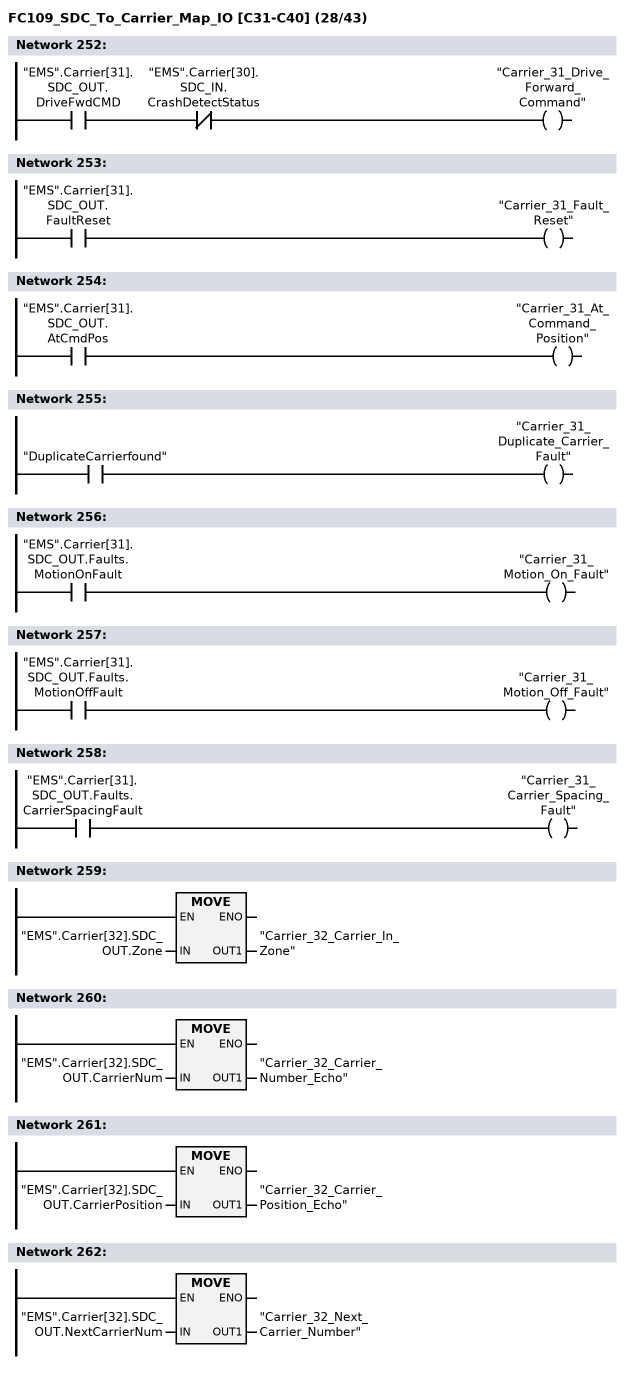
   RUNG wire#powerrail
      Contact( "EMS".Carrier[31].SDC_OUT.DriveFwdCMD )
      I_Contact( "EMS".Carrier[30].SDC_IN.CrashDetectStatus )
      Coil( "Carrier_31_Drive_Forward_Command" )
   END_RUNG
   // the same network as SCL:
   "Carrier_31_Drive_Forward_Command" := "EMS".Carrier[31].SDC_OUT.DriveFwdCMD AND NOT "EMS".Carrier[30].SDC_IN.CrashDetectStatus;
END_REGION

REGION Network 253
   RUNG wire#powerrail
      Contact( "EMS".Carrier[31].SDC_OUT.FaultReset )
      Coil( "Carrier_31_Fault_Reset" )
   END_RUNG
   // the same network as SCL:
   "Carrier_31_Fault_Reset" := "EMS".Carrier[31].SDC_OUT.FaultReset;
END_REGION

REGION Network 254
   RUNG wire#powerrail
      Contact( "EMS".Carrier[31].SDC_OUT.AtCmdPos )
      Coil( "Carrier_31_At_Command_Position" )
   END_RUNG
   // the same network as SCL:
   "Carrier_31_At_Command_Position" := "EMS".Carrier[31].SDC_OUT.AtCmdPos;
END_REGION

REGION Network 255
   RUNG wire#powerrail
      Contact( "DuplicateCarrierfound" )
      Coil( "Carrier_31_Duplicate_Carrier_Fault" )
   END_RUNG
   // the same network as SCL:
   "Carrier_31_Duplicate_Carrier_Fault" := "DuplicateCarrierfound";
END_REGION

REGION Network 256
   RUNG wire#powerrail
      Contact( "EMS".Carrier[31].SDC_OUT.Faults.MotionOnFault )
      Coil( "Carrier_31_Motion_On_Fault" )
   END_RUNG
   // the same network as SCL:
   "Carrier_31_Motion_On_Fault" := "EMS".Carrier[31].SDC_OUT.Faults.MotionOnFault;
END_REGION

REGION Network 257
   RUNG wire#powerrail
      Contact( "EMS".Carrier[31].SDC_OUT.Faults.MotionOffFault )
      Coil( "Carrier_31_Motion_Off_Fault" )
   END_RUNG
   // the same network as SCL:
   "Carrier_31_Motion_Off_Fault" := "EMS".Carrier[31].SDC_OUT.Faults.MotionOffFault;
END_REGION

REGION Network 258
   RUNG wire#powerrail
      Contact( "EMS".Carrier[31].SDC_OUT.Faults.CarrierSpacingFault )
      Coil( "Carrier_31_Carrier_Spacing_Fault" )
   END_RUNG
   // the same network as SCL:
   "Carrier_31_Carrier_Spacing_Fault" := "EMS".Carrier[31].SDC_OUT.Faults.CarrierSpacingFault;
END_REGION

REGION Network 259
   RUNG wire#powerrail
      Move(in := "EMS".Carrier[32].SDC_OUT.Zone, out1 => "Carrier_32_Carrier_In_Zone")
   END_RUNG
   // the same network as SCL:
   "Carrier_32_Carrier_In_Zone" := "EMS".Carrier[32].SDC_OUT.Zone;
END_REGION

REGION Network 260
   RUNG wire#powerrail
      Move(in := "EMS".Carrier[32].SDC_OUT.CarrierNum, out1 => "Carrier_32_Carrier_Number_Echo")
   END_RUNG
   // the same network as SCL:
   "Carrier_32_Carrier_Number_Echo" := "EMS".Carrier[32].SDC_OUT.CarrierNum;
END_REGION

REGION Network 261
   RUNG wire#powerrail
      Move(in := "EMS".Carrier[32].SDC_OUT.CarrierPosition, out1 => "Carrier_32_Carrier_Position_Echo")
   END_RUNG
   // the same network as SCL:
   "Carrier_32_Carrier_Position_Echo" := "EMS".Carrier[32].SDC_OUT.CarrierPosition;
END_REGION

REGION Network 262
   RUNG wire#powerrail
      Move(in := "EMS".Carrier[32].SDC_OUT.NextCarrierNum, out1 => "Carrier_32_Next_Carrier_Number")
   END_RUNG
   // the same network as SCL:
   "Carrier_32_Next_Carrier_Number" := "EMS".Carrier[32].SDC_OUT.NextCarrierNum;
END_REGION

REGION Network 263
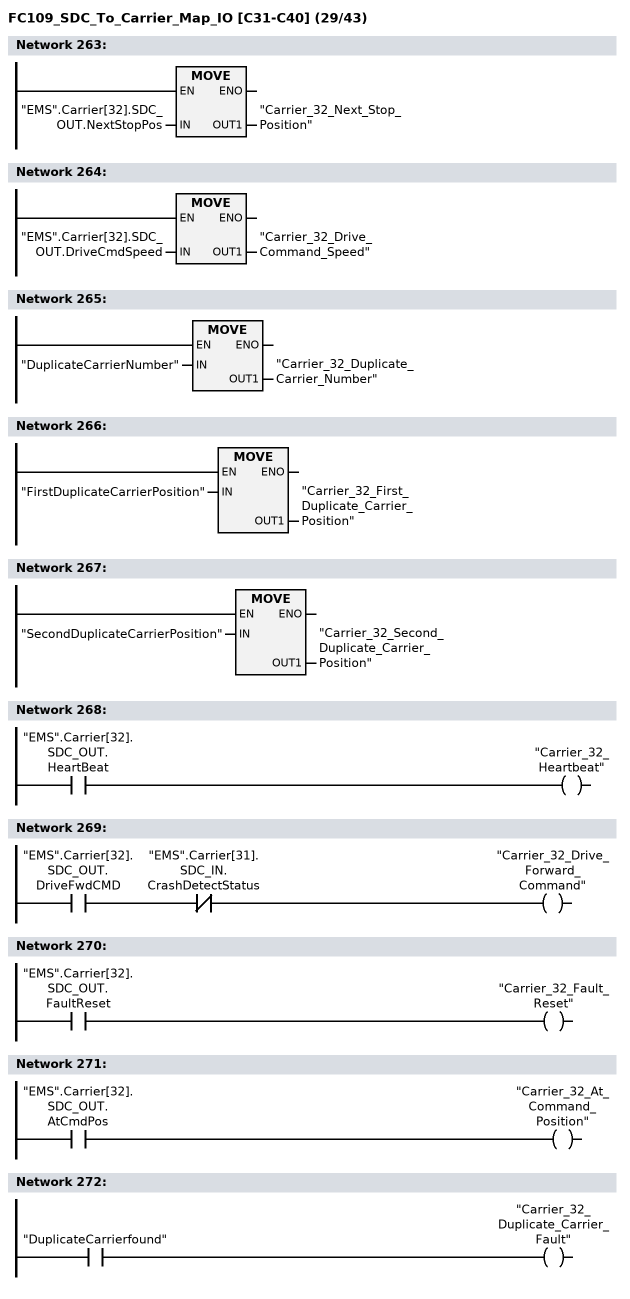
   RUNG wire#powerrail
      Move(in := "EMS".Carrier[32].SDC_OUT.NextStopPos, out1 => "Carrier_32_Next_Stop_Position")
   END_RUNG
   // the same network as SCL:
   "Carrier_32_Next_Stop_Position" := "EMS".Carrier[32].SDC_OUT.NextStopPos;
END_REGION

REGION Network 264
   RUNG wire#powerrail
      Move(in := "EMS".Carrier[32].SDC_OUT.DriveCmdSpeed, out1 => "Carrier_32_Drive_Command_Speed")
   END_RUNG
   // the same network as SCL:
   "Carrier_32_Drive_Command_Speed" := "EMS".Carrier[32].SDC_OUT.DriveCmdSpeed;
END_REGION

REGION Network 265
   RUNG wire#powerrail
      Move(in := "DuplicateCarrierNumber", out1 => "Carrier_32_Duplicate_Carrier_Number")
   END_RUNG
   // the same network as SCL:
   "Carrier_32_Duplicate_Carrier_Number" := "DuplicateCarrierNumber";
END_REGION

REGION Network 266
   RUNG wire#powerrail
      Move(in := "FirstDuplicateCarrierPosition", out1 => "Carrier_32_First_Duplicate_Carrier_Position")
   END_RUNG
   // the same network as SCL:
   "Carrier_32_First_Duplicate_Carrier_Position" := "FirstDuplicateCarrierPosition";
END_REGION

REGION Network 267
   RUNG wire#powerrail
      Move(in := "SecondDuplicateCarrierPosition", out1 => "Carrier_32_Second_Duplicate_Carrier_Position")
   END_RUNG
   // the same network as SCL:
   "Carrier_32_Second_Duplicate_Carrier_Position" := "SecondDuplicateCarrierPosition";
END_REGION

REGION Network 268
   RUNG wire#powerrail
      Contact( "EMS".Carrier[32].SDC_OUT.HeartBeat )
      Coil( "Carrier_32_Heartbeat" )
   END_RUNG
   // the same network as SCL:
   "Carrier_32_Heartbeat" := "EMS".Carrier[32].SDC_OUT.HeartBeat;
END_REGION

REGION Network 269
   RUNG wire#powerrail
      Contact( "EMS".Carrier[32].SDC_OUT.DriveFwdCMD )
      I_Contact( "EMS".Carrier[31].SDC_IN.CrashDetectStatus )
      Coil( "Carrier_32_Drive_Forward_Command" )
   END_RUNG
   // the same network as SCL:
   "Carrier_32_Drive_Forward_Command" := "EMS".Carrier[32].SDC_OUT.DriveFwdCMD AND NOT "EMS".Carrier[31].SDC_IN.CrashDetectStatus;
END_REGION

REGION Network 270
   RUNG wire#powerrail
      Contact( "EMS".Carrier[32].SDC_OUT.FaultReset )
      Coil( "Carrier_32_Fault_Reset" )
   END_RUNG
   // the same network as SCL:
   "Carrier_32_Fault_Reset" := "EMS".Carrier[32].SDC_OUT.FaultReset;
END_REGION

REGION Network 271
   RUNG wire#powerrail
      Contact( "EMS".Carrier[32].SDC_OUT.AtCmdPos )
      Coil( "Carrier_32_At_Command_Position" )
   END_RUNG
   // the same network as SCL:
   "Carrier_32_At_Command_Position" := "EMS".Carrier[32].SDC_OUT.AtCmdPos;
END_REGION

REGION Network 272
   RUNG wire#powerrail
      Contact( "DuplicateCarrierfound" )
      Coil( "Carrier_32_Duplicate_Carrier_Fault" )
   END_RUNG
   // the same network as SCL:
   "Carrier_32_Duplicate_Carrier_Fault" := "DuplicateCarrierfound";
END_REGION

REGION Network 273
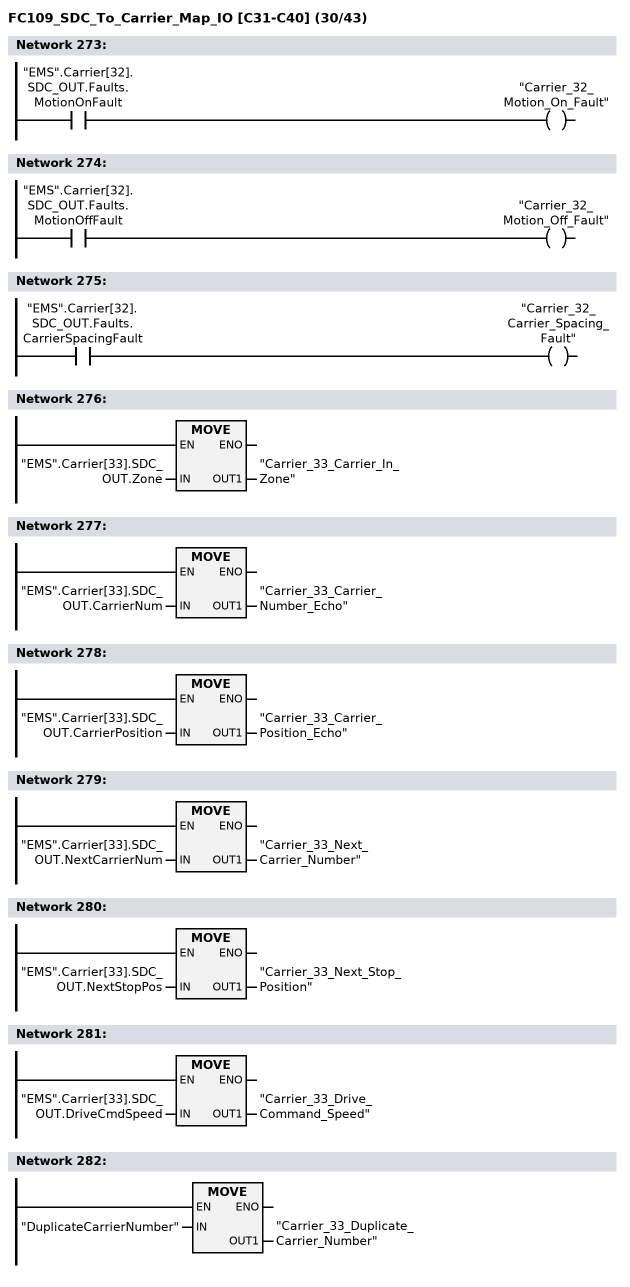
   RUNG wire#powerrail
      Contact( "EMS".Carrier[32].SDC_OUT.Faults.MotionOnFault )
      Coil( "Carrier_32_Motion_On_Fault" )
   END_RUNG
   // the same network as SCL:
   "Carrier_32_Motion_On_Fault" := "EMS".Carrier[32].SDC_OUT.Faults.MotionOnFault;
END_REGION

REGION Network 274
   RUNG wire#powerrail
      Contact( "EMS".Carrier[32].SDC_OUT.Faults.MotionOffFault )
      Coil( "Carrier_32_Motion_Off_Fault" )
   END_RUNG
   // the same network as SCL:
   "Carrier_32_Motion_Off_Fault" := "EMS".Carrier[32].SDC_OUT.Faults.MotionOffFault;
END_REGION

REGION Network 275
   RUNG wire#powerrail
      Contact( "EMS".Carrier[32].SDC_OUT.Faults.CarrierSpacingFault )
      Coil( "Carrier_32_Carrier_Spacing_Fault" )
   END_RUNG
   // the same network as SCL:
   "Carrier_32_Carrier_Spacing_Fault" := "EMS".Carrier[32].SDC_OUT.Faults.CarrierSpacingFault;
END_REGION

REGION Network 276
   RUNG wire#powerrail
      Move(in := "EMS".Carrier[33].SDC_OUT.Zone, out1 => "Carrier_33_Carrier_In_Zone")
   END_RUNG
   // the same network as SCL:
   "Carrier_33_Carrier_In_Zone" := "EMS".Carrier[33].SDC_OUT.Zone;
END_REGION

REGION Network 277
   RUNG wire#powerrail
      Move(in := "EMS".Carrier[33].SDC_OUT.CarrierNum, out1 => "Carrier_33_Carrier_Number_Echo")
   END_RUNG
   // the same network as SCL:
   "Carrier_33_Carrier_Number_Echo" := "EMS".Carrier[33].SDC_OUT.CarrierNum;
END_REGION

REGION Network 278
   RUNG wire#powerrail
      Move(in := "EMS".Carrier[33].SDC_OUT.CarrierPosition, out1 => "Carrier_33_Carrier_Position_Echo")
   END_RUNG
   // the same network as SCL:
   "Carrier_33_Carrier_Position_Echo" := "EMS".Carrier[33].SDC_OUT.CarrierPosition;
END_REGION

REGION Network 279
   RUNG wire#powerrail
      Move(in := "EMS".Carrier[33].SDC_OUT.NextCarrierNum, out1 => "Carrier_33_Next_Carrier_Number")
   END_RUNG
   // the same network as SCL:
   "Carrier_33_Next_Carrier_Number" := "EMS".Carrier[33].SDC_OUT.NextCarrierNum;
END_REGION

REGION Network 280
   RUNG wire#powerrail
      Move(in := "EMS".Carrier[33].SDC_OUT.NextStopPos, out1 => "Carrier_33_Next_Stop_Position")
   END_RUNG
   // the same network as SCL:
   "Carrier_33_Next_Stop_Position" := "EMS".Carrier[33].SDC_OUT.NextStopPos;
END_REGION

REGION Network 281
   RUNG wire#powerrail
      Move(in := "EMS".Carrier[33].SDC_OUT.DriveCmdSpeed, out1 => "Carrier_33_Drive_Command_Speed")
   END_RUNG
   // the same network as SCL:
   "Carrier_33_Drive_Command_Speed" := "EMS".Carrier[33].SDC_OUT.DriveCmdSpeed;
END_REGION

REGION Network 282
   RUNG wire#powerrail
      Move(in := "DuplicateCarrierNumber", out1 => "Carrier_33_Duplicate_Carrier_Number")
   END_RUNG
   // the same network as SCL:
   "Carrier_33_Duplicate_Carrier_Number" := "DuplicateCarrierNumber";
END_REGION

REGION Network 283
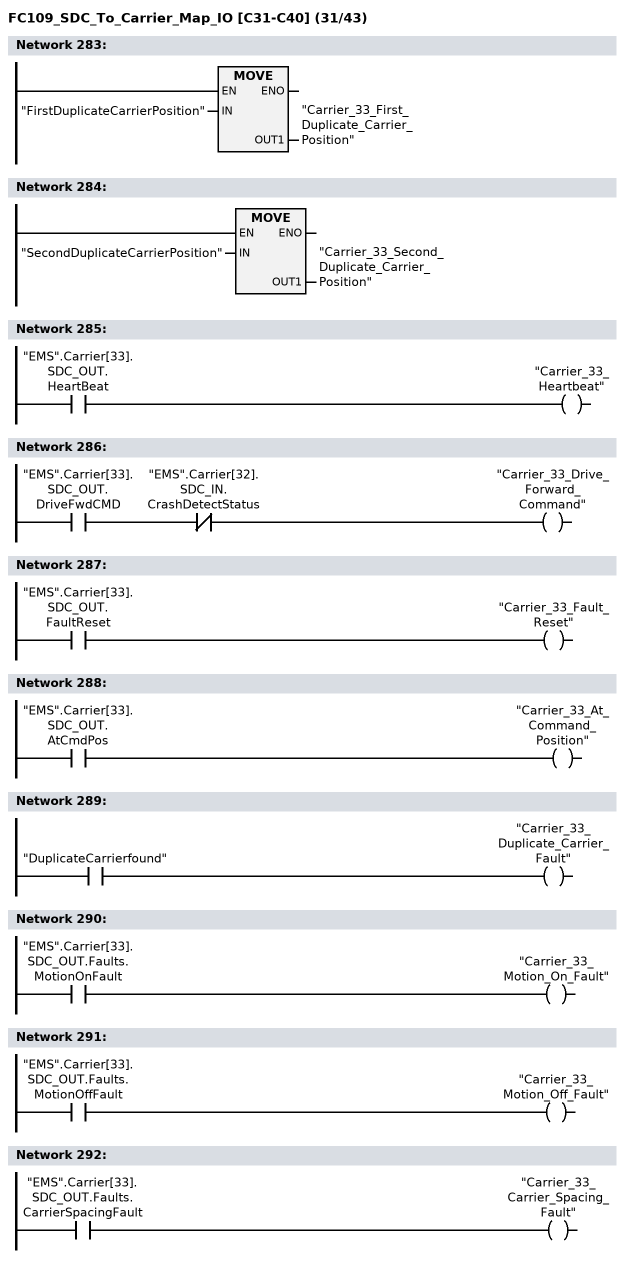
   RUNG wire#powerrail
      Move(in := "FirstDuplicateCarrierPosition", out1 => "Carrier_33_First_Duplicate_Carrier_Position")
   END_RUNG
   // the same network as SCL:
   "Carrier_33_First_Duplicate_Carrier_Position" := "FirstDuplicateCarrierPosition";
END_REGION

REGION Network 284
   RUNG wire#powerrail
      Move(in := "SecondDuplicateCarrierPosition", out1 => "Carrier_33_Second_Duplicate_Carrier_Position")
   END_RUNG
   // the same network as SCL:
   "Carrier_33_Second_Duplicate_Carrier_Position" := "SecondDuplicateCarrierPosition";
END_REGION

REGION Network 285
   RUNG wire#powerrail
      Contact( "EMS".Carrier[33].SDC_OUT.HeartBeat )
      Coil( "Carrier_33_Heartbeat" )
   END_RUNG
   // the same network as SCL:
   "Carrier_33_Heartbeat" := "EMS".Carrier[33].SDC_OUT.HeartBeat;
END_REGION

REGION Network 286
   RUNG wire#powerrail
      Contact( "EMS".Carrier[33].SDC_OUT.DriveFwdCMD )
      I_Contact( "EMS".Carrier[32].SDC_IN.CrashDetectStatus )
      Coil( "Carrier_33_Drive_Forward_Command" )
   END_RUNG
   // the same network as SCL:
   "Carrier_33_Drive_Forward_Command" := "EMS".Carrier[33].SDC_OUT.DriveFwdCMD AND NOT "EMS".Carrier[32].SDC_IN.CrashDetectStatus;
END_REGION

REGION Network 287
   RUNG wire#powerrail
      Contact( "EMS".Carrier[33].SDC_OUT.FaultReset )
      Coil( "Carrier_33_Fault_Reset" )
   END_RUNG
   // the same network as SCL:
   "Carrier_33_Fault_Reset" := "EMS".Carrier[33].SDC_OUT.FaultReset;
END_REGION

REGION Network 288
   RUNG wire#powerrail
      Contact( "EMS".Carrier[33].SDC_OUT.AtCmdPos )
      Coil( "Carrier_33_At_Command_Position" )
   END_RUNG
   // the same network as SCL:
   "Carrier_33_At_Command_Position" := "EMS".Carrier[33].SDC_OUT.AtCmdPos;
END_REGION

REGION Network 289
   RUNG wire#powerrail
      Contact( "DuplicateCarrierfound" )
      Coil( "Carrier_33_Duplicate_Carrier_Fault" )
   END_RUNG
   // the same network as SCL:
   "Carrier_33_Duplicate_Carrier_Fault" := "DuplicateCarrierfound";
END_REGION

REGION Network 290
   RUNG wire#powerrail
      Contact( "EMS".Carrier[33].SDC_OUT.Faults.MotionOnFault )
      Coil( "Carrier_33_Motion_On_Fault" )
   END_RUNG
   // the same network as SCL:
   "Carrier_33_Motion_On_Fault" := "EMS".Carrier[33].SDC_OUT.Faults.MotionOnFault;
END_REGION

REGION Network 291
   RUNG wire#powerrail
      Contact( "EMS".Carrier[33].SDC_OUT.Faults.MotionOffFault )
      Coil( "Carrier_33_Motion_Off_Fault" )
   END_RUNG
   // the same network as SCL:
   "Carrier_33_Motion_Off_Fault" := "EMS".Carrier[33].SDC_OUT.Faults.MotionOffFault;
END_REGION

REGION Network 292
   RUNG wire#powerrail
      Contact( "EMS".Carrier[33].SDC_OUT.Faults.CarrierSpacingFault )
      Coil( "Carrier_33_Carrier_Spacing_Fault" )
   END_RUNG
   // the same network as SCL:
   "Carrier_33_Carrier_Spacing_Fault" := "EMS".Carrier[33].SDC_OUT.Faults.CarrierSpacingFault;
END_REGION

REGION Network 293
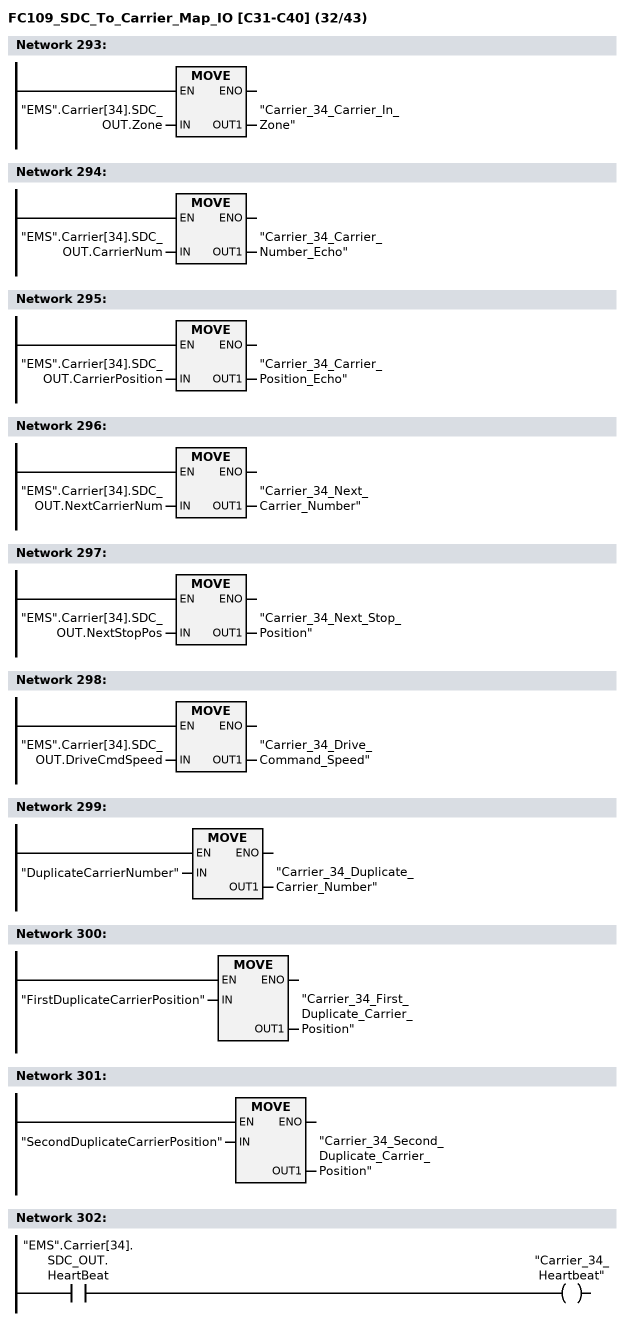
   RUNG wire#powerrail
      Move(in := "EMS".Carrier[34].SDC_OUT.Zone, out1 => "Carrier_34_Carrier_In_Zone")
   END_RUNG
   // the same network as SCL:
   "Carrier_34_Carrier_In_Zone" := "EMS".Carrier[34].SDC_OUT.Zone;
END_REGION

REGION Network 294
   RUNG wire#powerrail
      Move(in := "EMS".Carrier[34].SDC_OUT.CarrierNum, out1 => "Carrier_34_Carrier_Number_Echo")
   END_RUNG
   // the same network as SCL:
   "Carrier_34_Carrier_Number_Echo" := "EMS".Carrier[34].SDC_OUT.CarrierNum;
END_REGION

REGION Network 295
   RUNG wire#powerrail
      Move(in := "EMS".Carrier[34].SDC_OUT.CarrierPosition, out1 => "Carrier_34_Carrier_Position_Echo")
   END_RUNG
   // the same network as SCL:
   "Carrier_34_Carrier_Position_Echo" := "EMS".Carrier[34].SDC_OUT.CarrierPosition;
END_REGION

REGION Network 296
   RUNG wire#powerrail
      Move(in := "EMS".Carrier[34].SDC_OUT.NextCarrierNum, out1 => "Carrier_34_Next_Carrier_Number")
   END_RUNG
   // the same network as SCL:
   "Carrier_34_Next_Carrier_Number" := "EMS".Carrier[34].SDC_OUT.NextCarrierNum;
END_REGION

REGION Network 297
   RUNG wire#powerrail
      Move(in := "EMS".Carrier[34].SDC_OUT.NextStopPos, out1 => "Carrier_34_Next_Stop_Position")
   END_RUNG
   // the same network as SCL:
   "Carrier_34_Next_Stop_Position" := "EMS".Carrier[34].SDC_OUT.NextStopPos;
END_REGION

REGION Network 298
   RUNG wire#powerrail
      Move(in := "EMS".Carrier[34].SDC_OUT.DriveCmdSpeed, out1 => "Carrier_34_Drive_Command_Speed")
   END_RUNG
   // the same network as SCL:
   "Carrier_34_Drive_Command_Speed" := "EMS".Carrier[34].SDC_OUT.DriveCmdSpeed;
END_REGION

REGION Network 299
   RUNG wire#powerrail
      Move(in := "DuplicateCarrierNumber", out1 => "Carrier_34_Duplicate_Carrier_Number")
   END_RUNG
   // the same network as SCL:
   "Carrier_34_Duplicate_Carrier_Number" := "DuplicateCarrierNumber";
END_REGION

REGION Network 300
   RUNG wire#powerrail
      Move(in := "FirstDuplicateCarrierPosition", out1 => "Carrier_34_First_Duplicate_Carrier_Position")
   END_RUNG
   // the same network as SCL:
   "Carrier_34_First_Duplicate_Carrier_Position" := "FirstDuplicateCarrierPosition";
END_REGION

REGION Network 301
   RUNG wire#powerrail
      Move(in := "SecondDuplicateCarrierPosition", out1 => "Carrier_34_Second_Duplicate_Carrier_Position")
   END_RUNG
   // the same network as SCL:
   "Carrier_34_Second_Duplicate_Carrier_Position" := "SecondDuplicateCarrierPosition";
END_REGION

REGION Network 302
   RUNG wire#powerrail
      Contact( "EMS".Carrier[34].SDC_OUT.HeartBeat )
      Coil( "Carrier_34_Heartbeat" )
   END_RUNG
   // the same network as SCL:
   "Carrier_34_Heartbeat" := "EMS".Carrier[34].SDC_OUT.HeartBeat;
END_REGION

REGION Network 303
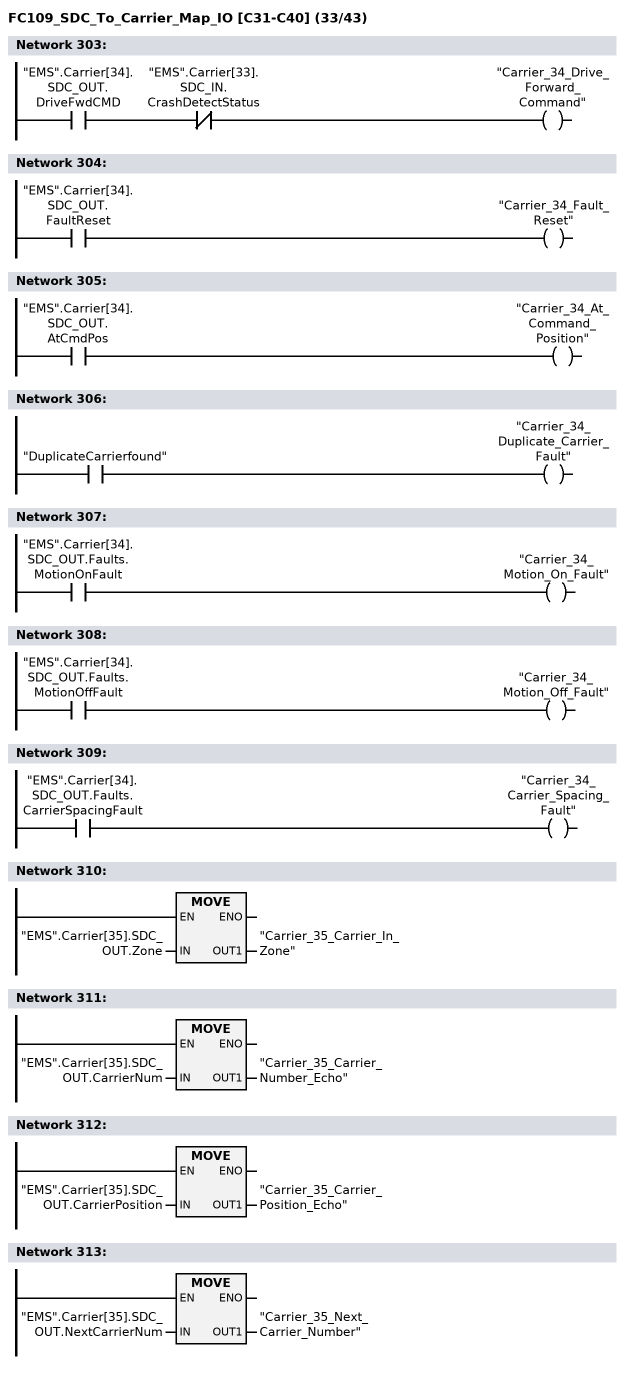
   RUNG wire#powerrail
      Contact( "EMS".Carrier[34].SDC_OUT.DriveFwdCMD )
      I_Contact( "EMS".Carrier[33].SDC_IN.CrashDetectStatus )
      Coil( "Carrier_34_Drive_Forward_Command" )
   END_RUNG
   // the same network as SCL:
   "Carrier_34_Drive_Forward_Command" := "EMS".Carrier[34].SDC_OUT.DriveFwdCMD AND NOT "EMS".Carrier[33].SDC_IN.CrashDetectStatus;
END_REGION

REGION Network 304
   RUNG wire#powerrail
      Contact( "EMS".Carrier[34].SDC_OUT.FaultReset )
      Coil( "Carrier_34_Fault_Reset" )
   END_RUNG
   // the same network as SCL:
   "Carrier_34_Fault_Reset" := "EMS".Carrier[34].SDC_OUT.FaultReset;
END_REGION

REGION Network 305
   RUNG wire#powerrail
      Contact( "EMS".Carrier[34].SDC_OUT.AtCmdPos )
      Coil( "Carrier_34_At_Command_Position" )
   END_RUNG
   // the same network as SCL:
   "Carrier_34_At_Command_Position" := "EMS".Carrier[34].SDC_OUT.AtCmdPos;
END_REGION

REGION Network 306
   RUNG wire#powerrail
      Contact( "DuplicateCarrierfound" )
      Coil( "Carrier_34_Duplicate_Carrier_Fault" )
   END_RUNG
   // the same network as SCL:
   "Carrier_34_Duplicate_Carrier_Fault" := "DuplicateCarrierfound";
END_REGION

REGION Network 307
   RUNG wire#powerrail
      Contact( "EMS".Carrier[34].SDC_OUT.Faults.MotionOnFault )
      Coil( "Carrier_34_Motion_On_Fault" )
   END_RUNG
   // the same network as SCL:
   "Carrier_34_Motion_On_Fault" := "EMS".Carrier[34].SDC_OUT.Faults.MotionOnFault;
END_REGION

REGION Network 308
   RUNG wire#powerrail
      Contact( "EMS".Carrier[34].SDC_OUT.Faults.MotionOffFault )
      Coil( "Carrier_34_Motion_Off_Fault" )
   END_RUNG
   // the same network as SCL:
   "Carrier_34_Motion_Off_Fault" := "EMS".Carrier[34].SDC_OUT.Faults.MotionOffFault;
END_REGION

REGION Network 309
   RUNG wire#powerrail
      Contact( "EMS".Carrier[34].SDC_OUT.Faults.CarrierSpacingFault )
      Coil( "Carrier_34_Carrier_Spacing_Fault" )
   END_RUNG
   // the same network as SCL:
   "Carrier_34_Carrier_Spacing_Fault" := "EMS".Carrier[34].SDC_OUT.Faults.CarrierSpacingFault;
END_REGION

REGION Network 310
   RUNG wire#powerrail
      Move(in := "EMS".Carrier[35].SDC_OUT.Zone, out1 => "Carrier_35_Carrier_In_Zone")
   END_RUNG
   // the same network as SCL:
   "Carrier_35_Carrier_In_Zone" := "EMS".Carrier[35].SDC_OUT.Zone;
END_REGION

REGION Network 311
   RUNG wire#powerrail
      Move(in := "EMS".Carrier[35].SDC_OUT.CarrierNum, out1 => "Carrier_35_Carrier_Number_Echo")
   END_RUNG
   // the same network as SCL:
   "Carrier_35_Carrier_Number_Echo" := "EMS".Carrier[35].SDC_OUT.CarrierNum;
END_REGION

REGION Network 312
   RUNG wire#powerrail
      Move(in := "EMS".Carrier[35].SDC_OUT.CarrierPosition, out1 => "Carrier_35_Carrier_Position_Echo")
   END_RUNG
   // the same network as SCL:
   "Carrier_35_Carrier_Position_Echo" := "EMS".Carrier[35].SDC_OUT.CarrierPosition;
END_REGION

REGION Network 313
   RUNG wire#powerrail
      Move(in := "EMS".Carrier[35].SDC_OUT.NextCarrierNum, out1 => "Carrier_35_Next_Carrier_Number")
   END_RUNG
   // the same network as SCL:
   "Carrier_35_Next_Carrier_Number" := "EMS".Carrier[35].SDC_OUT.NextCarrierNum;
END_REGION

REGION Network 314
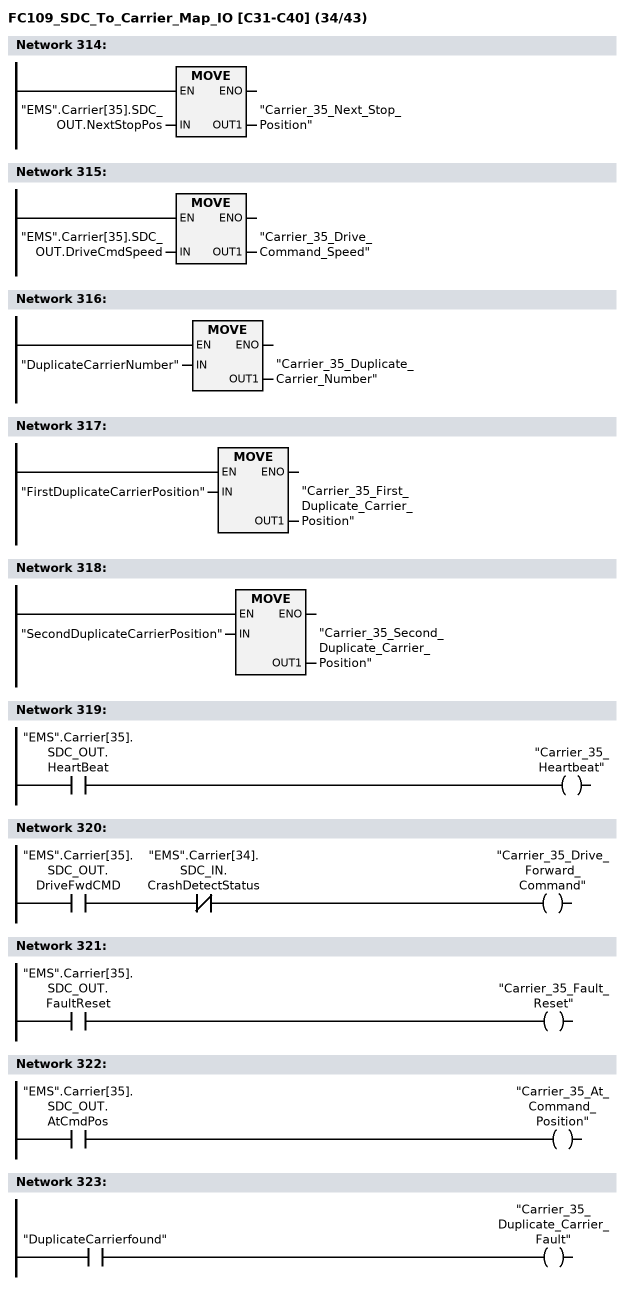
   RUNG wire#powerrail
      Move(in := "EMS".Carrier[35].SDC_OUT.NextStopPos, out1 => "Carrier_35_Next_Stop_Position")
   END_RUNG
   // the same network as SCL:
   "Carrier_35_Next_Stop_Position" := "EMS".Carrier[35].SDC_OUT.NextStopPos;
END_REGION

REGION Network 315
   RUNG wire#powerrail
      Move(in := "EMS".Carrier[35].SDC_OUT.DriveCmdSpeed, out1 => "Carrier_35_Drive_Command_Speed")
   END_RUNG
   // the same network as SCL:
   "Carrier_35_Drive_Command_Speed" := "EMS".Carrier[35].SDC_OUT.DriveCmdSpeed;
END_REGION

REGION Network 316
   RUNG wire#powerrail
      Move(in := "DuplicateCarrierNumber", out1 => "Carrier_35_Duplicate_Carrier_Number")
   END_RUNG
   // the same network as SCL:
   "Carrier_35_Duplicate_Carrier_Number" := "DuplicateCarrierNumber";
END_REGION

REGION Network 317
   RUNG wire#powerrail
      Move(in := "FirstDuplicateCarrierPosition", out1 => "Carrier_35_First_Duplicate_Carrier_Position")
   END_RUNG
   // the same network as SCL:
   "Carrier_35_First_Duplicate_Carrier_Position" := "FirstDuplicateCarrierPosition";
END_REGION

REGION Network 318
   RUNG wire#powerrail
      Move(in := "SecondDuplicateCarrierPosition", out1 => "Carrier_35_Second_Duplicate_Carrier_Position")
   END_RUNG
   // the same network as SCL:
   "Carrier_35_Second_Duplicate_Carrier_Position" := "SecondDuplicateCarrierPosition";
END_REGION

REGION Network 319
   RUNG wire#powerrail
      Contact( "EMS".Carrier[35].SDC_OUT.HeartBeat )
      Coil( "Carrier_35_Heartbeat" )
   END_RUNG
   // the same network as SCL:
   "Carrier_35_Heartbeat" := "EMS".Carrier[35].SDC_OUT.HeartBeat;
END_REGION

REGION Network 320
   RUNG wire#powerrail
      Contact( "EMS".Carrier[35].SDC_OUT.DriveFwdCMD )
      I_Contact( "EMS".Carrier[34].SDC_IN.CrashDetectStatus )
      Coil( "Carrier_35_Drive_Forward_Command" )
   END_RUNG
   // the same network as SCL:
   "Carrier_35_Drive_Forward_Command" := "EMS".Carrier[35].SDC_OUT.DriveFwdCMD AND NOT "EMS".Carrier[34].SDC_IN.CrashDetectStatus;
END_REGION

REGION Network 321
   RUNG wire#powerrail
      Contact( "EMS".Carrier[35].SDC_OUT.FaultReset )
      Coil( "Carrier_35_Fault_Reset" )
   END_RUNG
   // the same network as SCL:
   "Carrier_35_Fault_Reset" := "EMS".Carrier[35].SDC_OUT.FaultReset;
END_REGION

REGION Network 322
   RUNG wire#powerrail
      Contact( "EMS".Carrier[35].SDC_OUT.AtCmdPos )
      Coil( "Carrier_35_At_Command_Position" )
   END_RUNG
   // the same network as SCL:
   "Carrier_35_At_Command_Position" := "EMS".Carrier[35].SDC_OUT.AtCmdPos;
END_REGION

REGION Network 323
   RUNG wire#powerrail
      Contact( "DuplicateCarrierfound" )
      Coil( "Carrier_35_Duplicate_Carrier_Fault" )
   END_RUNG
   // the same network as SCL:
   "Carrier_35_Duplicate_Carrier_Fault" := "DuplicateCarrierfound";
END_REGION

REGION Network 324
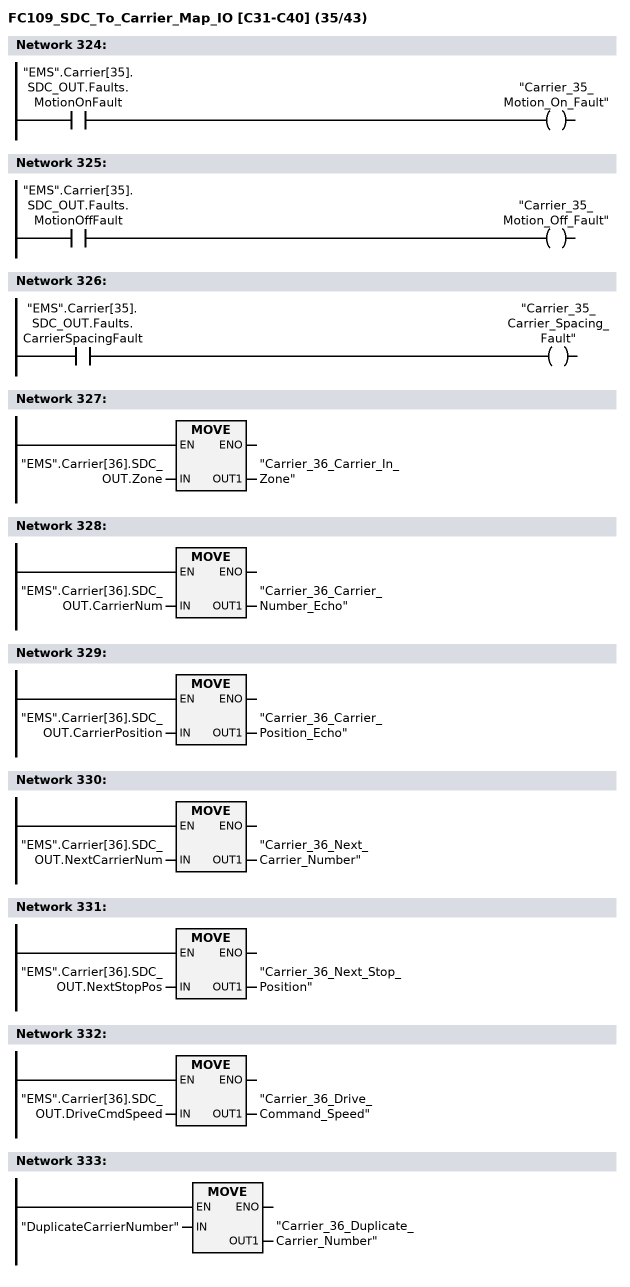
   RUNG wire#powerrail
      Contact( "EMS".Carrier[35].SDC_OUT.Faults.MotionOnFault )
      Coil( "Carrier_35_Motion_On_Fault" )
   END_RUNG
   // the same network as SCL:
   "Carrier_35_Motion_On_Fault" := "EMS".Carrier[35].SDC_OUT.Faults.MotionOnFault;
END_REGION

REGION Network 325
   RUNG wire#powerrail
      Contact( "EMS".Carrier[35].SDC_OUT.Faults.MotionOffFault )
      Coil( "Carrier_35_Motion_Off_Fault" )
   END_RUNG
   // the same network as SCL:
   "Carrier_35_Motion_Off_Fault" := "EMS".Carrier[35].SDC_OUT.Faults.MotionOffFault;
END_REGION

REGION Network 326
   RUNG wire#powerrail
      Contact( "EMS".Carrier[35].SDC_OUT.Faults.CarrierSpacingFault )
      Coil( "Carrier_35_Carrier_Spacing_Fault" )
   END_RUNG
   // the same network as SCL:
   "Carrier_35_Carrier_Spacing_Fault" := "EMS".Carrier[35].SDC_OUT.Faults.CarrierSpacingFault;
END_REGION

REGION Network 327
   RUNG wire#powerrail
      Move(in := "EMS".Carrier[36].SDC_OUT.Zone, out1 => "Carrier_36_Carrier_In_Zone")
   END_RUNG
   // the same network as SCL:
   "Carrier_36_Carrier_In_Zone" := "EMS".Carrier[36].SDC_OUT.Zone;
END_REGION

REGION Network 328
   RUNG wire#powerrail
      Move(in := "EMS".Carrier[36].SDC_OUT.CarrierNum, out1 => "Carrier_36_Carrier_Number_Echo")
   END_RUNG
   // the same network as SCL:
   "Carrier_36_Carrier_Number_Echo" := "EMS".Carrier[36].SDC_OUT.CarrierNum;
END_REGION

REGION Network 329
   RUNG wire#powerrail
      Move(in := "EMS".Carrier[36].SDC_OUT.CarrierPosition, out1 => "Carrier_36_Carrier_Position_Echo")
   END_RUNG
   // the same network as SCL:
   "Carrier_36_Carrier_Position_Echo" := "EMS".Carrier[36].SDC_OUT.CarrierPosition;
END_REGION

REGION Network 330
   RUNG wire#powerrail
      Move(in := "EMS".Carrier[36].SDC_OUT.NextCarrierNum, out1 => "Carrier_36_Next_Carrier_Number")
   END_RUNG
   // the same network as SCL:
   "Carrier_36_Next_Carrier_Number" := "EMS".Carrier[36].SDC_OUT.NextCarrierNum;
END_REGION

REGION Network 331
   RUNG wire#powerrail
      Move(in := "EMS".Carrier[36].SDC_OUT.NextStopPos, out1 => "Carrier_36_Next_Stop_Position")
   END_RUNG
   // the same network as SCL:
   "Carrier_36_Next_Stop_Position" := "EMS".Carrier[36].SDC_OUT.NextStopPos;
END_REGION

REGION Network 332
   RUNG wire#powerrail
      Move(in := "EMS".Carrier[36].SDC_OUT.DriveCmdSpeed, out1 => "Carrier_36_Drive_Command_Speed")
   END_RUNG
   // the same network as SCL:
   "Carrier_36_Drive_Command_Speed" := "EMS".Carrier[36].SDC_OUT.DriveCmdSpeed;
END_REGION

REGION Network 333
   RUNG wire#powerrail
      Move(in := "DuplicateCarrierNumber", out1 => "Carrier_36_Duplicate_Carrier_Number")
   END_RUNG
   // the same network as SCL:
   "Carrier_36_Duplicate_Carrier_Number" := "DuplicateCarrierNumber";
END_REGION

REGION Network 334
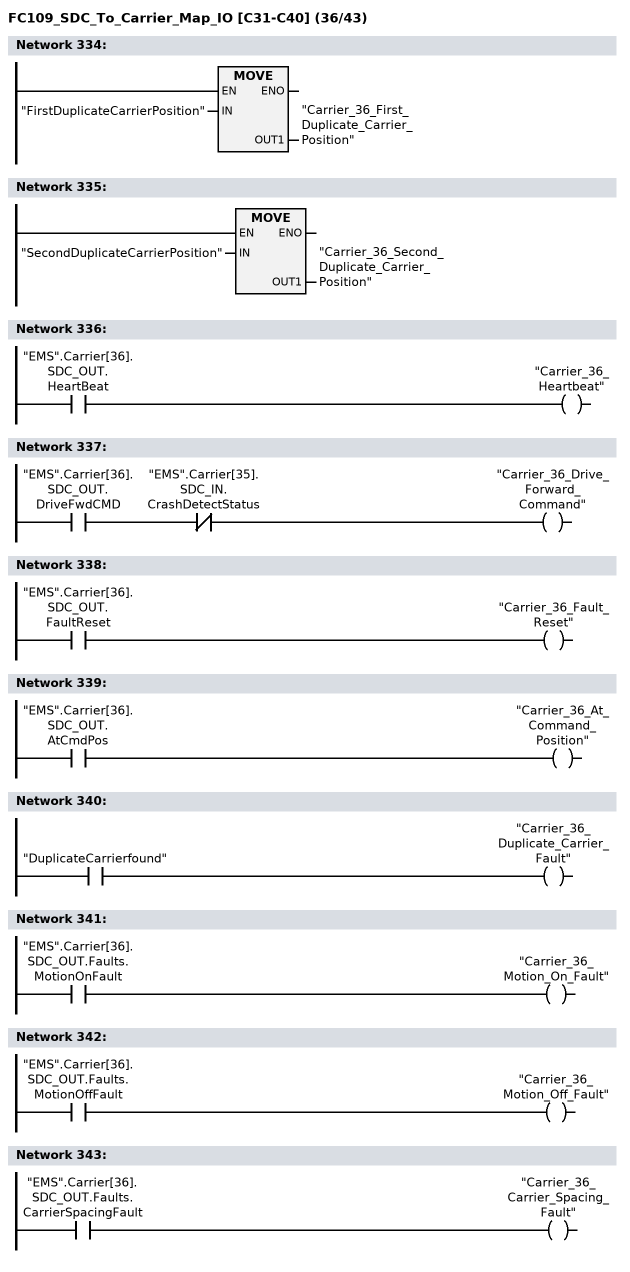
   RUNG wire#powerrail
      Move(in := "FirstDuplicateCarrierPosition", out1 => "Carrier_36_First_Duplicate_Carrier_Position")
   END_RUNG
   // the same network as SCL:
   "Carrier_36_First_Duplicate_Carrier_Position" := "FirstDuplicateCarrierPosition";
END_REGION

REGION Network 335
   RUNG wire#powerrail
      Move(in := "SecondDuplicateCarrierPosition", out1 => "Carrier_36_Second_Duplicate_Carrier_Position")
   END_RUNG
   // the same network as SCL:
   "Carrier_36_Second_Duplicate_Carrier_Position" := "SecondDuplicateCarrierPosition";
END_REGION

REGION Network 336
   RUNG wire#powerrail
      Contact( "EMS".Carrier[36].SDC_OUT.HeartBeat )
      Coil( "Carrier_36_Heartbeat" )
   END_RUNG
   // the same network as SCL:
   "Carrier_36_Heartbeat" := "EMS".Carrier[36].SDC_OUT.HeartBeat;
END_REGION

REGION Network 337
   RUNG wire#powerrail
      Contact( "EMS".Carrier[36].SDC_OUT.DriveFwdCMD )
      I_Contact( "EMS".Carrier[35].SDC_IN.CrashDetectStatus )
      Coil( "Carrier_36_Drive_Forward_Command" )
   END_RUNG
   // the same network as SCL:
   "Carrier_36_Drive_Forward_Command" := "EMS".Carrier[36].SDC_OUT.DriveFwdCMD AND NOT "EMS".Carrier[35].SDC_IN.CrashDetectStatus;
END_REGION

REGION Network 338
   RUNG wire#powerrail
      Contact( "EMS".Carrier[36].SDC_OUT.FaultReset )
      Coil( "Carrier_36_Fault_Reset" )
   END_RUNG
   // the same network as SCL:
   "Carrier_36_Fault_Reset" := "EMS".Carrier[36].SDC_OUT.FaultReset;
END_REGION

REGION Network 339
   RUNG wire#powerrail
      Contact( "EMS".Carrier[36].SDC_OUT.AtCmdPos )
      Coil( "Carrier_36_At_Command_Position" )
   END_RUNG
   // the same network as SCL:
   "Carrier_36_At_Command_Position" := "EMS".Carrier[36].SDC_OUT.AtCmdPos;
END_REGION

REGION Network 340
   RUNG wire#powerrail
      Contact( "DuplicateCarrierfound" )
      Coil( "Carrier_36_Duplicate_Carrier_Fault" )
   END_RUNG
   // the same network as SCL:
   "Carrier_36_Duplicate_Carrier_Fault" := "DuplicateCarrierfound";
END_REGION

REGION Network 341
   RUNG wire#powerrail
      Contact( "EMS".Carrier[36].SDC_OUT.Faults.MotionOnFault )
      Coil( "Carrier_36_Motion_On_Fault" )
   END_RUNG
   // the same network as SCL:
   "Carrier_36_Motion_On_Fault" := "EMS".Carrier[36].SDC_OUT.Faults.MotionOnFault;
END_REGION

REGION Network 342
   RUNG wire#powerrail
      Contact( "EMS".Carrier[36].SDC_OUT.Faults.MotionOffFault )
      Coil( "Carrier_36_Motion_Off_Fault" )
   END_RUNG
   // the same network as SCL:
   "Carrier_36_Motion_Off_Fault" := "EMS".Carrier[36].SDC_OUT.Faults.MotionOffFault;
END_REGION

REGION Network 343
   RUNG wire#powerrail
      Contact( "EMS".Carrier[36].SDC_OUT.Faults.CarrierSpacingFault )
      Coil( "Carrier_36_Carrier_Spacing_Fault" )
   END_RUNG
   // the same network as SCL:
   "Carrier_36_Carrier_Spacing_Fault" := "EMS".Carrier[36].SDC_OUT.Faults.CarrierSpacingFault;
END_REGION

REGION Network 344
